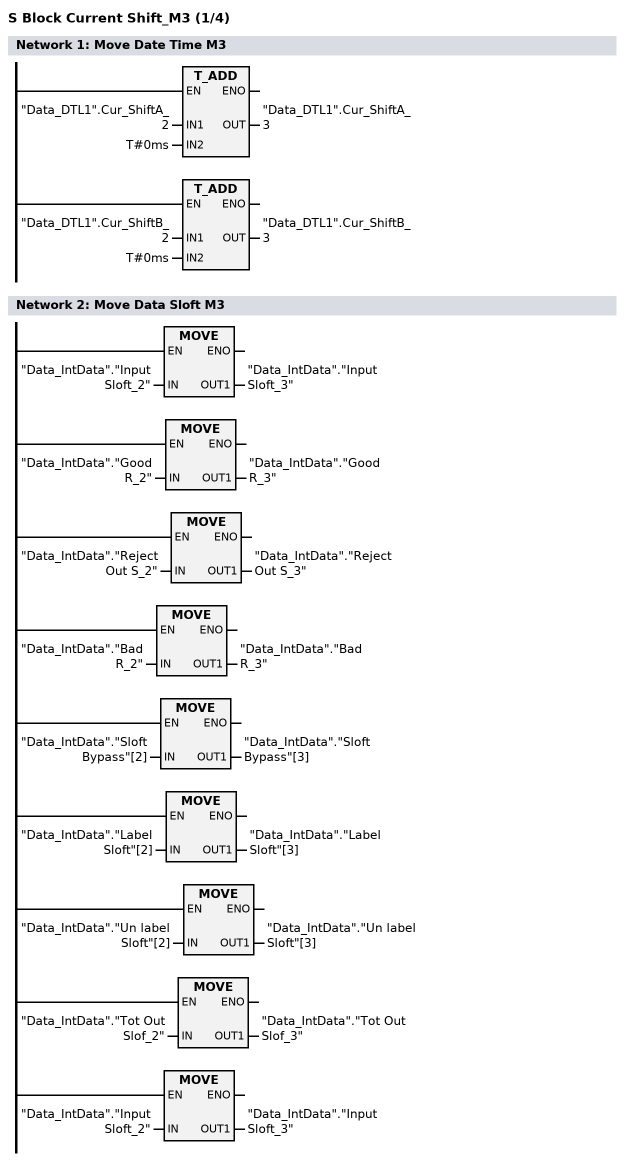
   "Data_DTL1".Cur_ShiftA_3 := T_ADD(IN1 := "Data_DTL1".Cur_ShiftA_2, IN2 := T#0ms);
   "Data_DTL1".Cur_ShiftB_3 := T_ADD(IN1 := "Data_DTL1".Cur_ShiftB_2, IN2 := T#0ms);
END_REGION

REGION Network 2: Move Data Sloft M3
   RUNG wire#powerrail
      { S7_GenerateENO := "TRUE" } Move(in := "Data_IntData"."Input Sloft_2", out1 => "Data_IntData"."Input Sloft_3")
   END_RUNG
   RUNG wire#powerrail
      { S7_GenerateENO := "TRUE" } Move(in := "Data_IntData"."Good R_2", out1 => "Data_IntData"."Good R_3")
   END_RUNG
   RUNG wire#powerrail
      { S7_GenerateENO := "TRUE" } Move(in := "Data_IntData"."Reject Out S_2", out1 => "Data_IntData"."Reject Out S_3")
   END_RUNG
   RUNG wire#powerrail
      { S7_GenerateENO := "TRUE" } Move(in := "Data_IntData"."Bad R_2", out1 => "Data_IntData"."Bad R_3")
   END_RUNG
   RUNG wire#powerrail
      { S7_GenerateENO := "TRUE" } Move(in := "Data_IntData"."Sloft Bypass"[2], out1 => "Data_IntData"."Sloft Bypass"[3])
   END_RUNG
   RUNG wire#powerrail
      { S7_GenerateENO := "TRUE" } Move(in := "Data_IntData"."Label Sloft"[2], out1 => "Data_IntData"."Label Sloft"[3])
   END_RUNG
   RUNG wire#powerrail
      { S7_GenerateENO := "TRUE" } Move(in := "Data_IntData"."Un label Sloft"[2], out1 => "Data_IntData"."Un label Sloft"[3])
   END_RUNG
   RUNG wire#powerrail
      { S7_GenerateENO := "TRUE" } Move(in := "Data_IntData"."Tot Out Slof_2", out1 => "Data_IntData"."Tot Out Slof_3")
   END_RUNG
   RUNG wire#powerrail
      { S7_GenerateENO := "TRUE" } Move(in := "Data_IntData"."Input Sloft_2", out1 => "Data_IntData"."Input Sloft_3")
   END_RUNG
   // the same network as SCL:
   "Data_IntData"."Input Sloft_3" := "Data_IntData"."Input Sloft_2";
   "Data_IntData"."Good R_3" := "Data_IntData"."Good R_2";
   "Data_IntData"."Reject Out S_3" := "Data_IntData"."Reject Out S_2";
   "Data_IntData"."Bad R_3" := "Data_IntData"."Bad R_2";
   "Data_IntData"."Sloft Bypass"[3] := "Data_IntData"."Sloft Bypass"[2];
   "Data_IntData"."Label Sloft"[3] := "Data_IntData"."Label Sloft"[2];
   "Data_IntData"."Un label Sloft"[3] := "Data_IntData"."Un label Sloft"[2];
   "Data_IntData"."Tot Out Slof_3" := "Data_IntData"."Tot Out Slof_2";
   "Data_IntData"."Input Sloft_3" := "Data_IntData"."Input Sloft_2";
END_REGION

REGION Network 3: Move Data Sloft Trigger & Aplicator M3
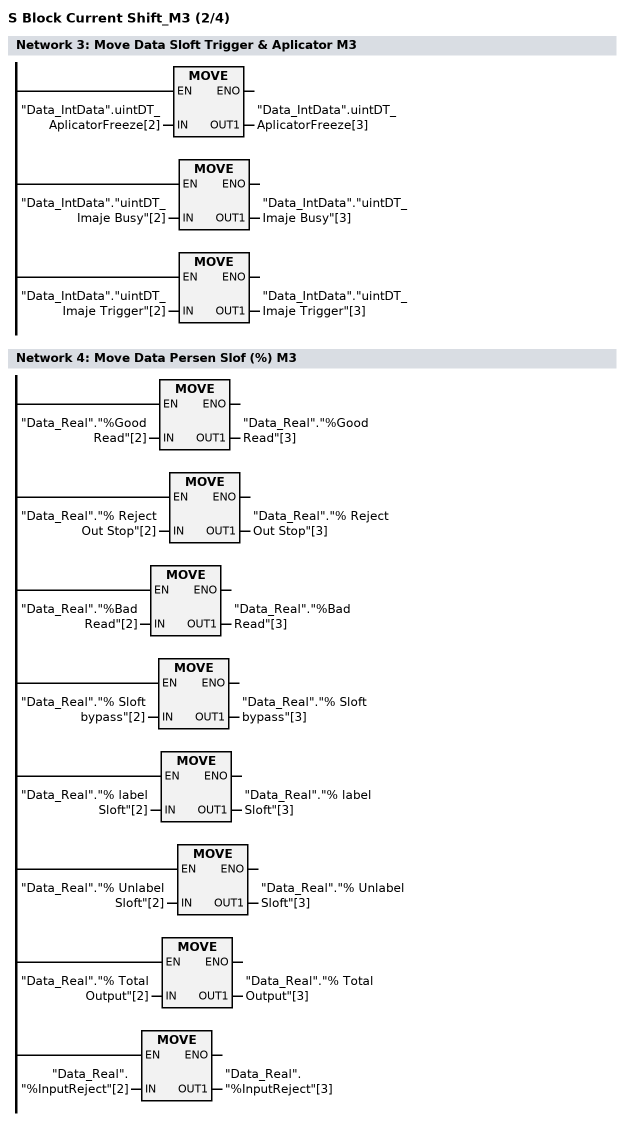
   RUNG wire#powerrail
      { S7_GenerateENO := "TRUE" } Move(in := "Data_IntData".uintDT_AplicatorFreeze[2], out1 => "Data_IntData".uintDT_AplicatorFreeze[3])
   END_RUNG
   RUNG wire#powerrail
      { S7_GenerateENO := "TRUE" } Move(in := "Data_IntData"."uintDT_Imaje Busy"[2], out1 => "Data_IntData"."uintDT_Imaje Busy"[3])
   END_RUNG
   RUNG wire#powerrail
      { S7_GenerateENO := "TRUE" } Move(in := "Data_IntData"."uintDT_Imaje Trigger"[2], out1 => "Data_IntData"."uintDT_Imaje Trigger"[3])
   END_RUNG
   // the same network as SCL:
   "Data_IntData".uintDT_AplicatorFreeze[3] := "Data_IntData".uintDT_AplicatorFreeze[2];
   "Data_IntData"."uintDT_Imaje Busy"[3] := "Data_IntData"."uintDT_Imaje Busy"[2];
   "Data_IntData"."uintDT_Imaje Trigger"[3] := "Data_IntData"."uintDT_Imaje Trigger"[2];
END_REGION

REGION Network 4: Move Data Persen Slof (%) M3
   RUNG wire#powerrail
      { S7_GenerateENO := "TRUE" } Move(in := "Data_Real"."%Good Read"[2], out1 => "Data_Real"."%Good Read"[3])
   END_RUNG
   RUNG wire#powerrail
      { S7_GenerateENO := "TRUE" } Move(in := "Data_Real"."% Reject Out Stop"[2], out1 => "Data_Real"."% Reject Out Stop"[3])
   END_RUNG
   RUNG wire#powerrail
      { S7_GenerateENO := "TRUE" } Move(in := "Data_Real"."%Bad Read"[2], out1 => "Data_Real"."%Bad Read"[3])
   END_RUNG
   RUNG wire#powerrail
      { S7_GenerateENO := "TRUE" } Move(in := "Data_Real"."% Sloft bypass"[2], out1 => "Data_Real"."% Sloft bypass"[3])
   END_RUNG
   RUNG wire#powerrail
      { S7_GenerateENO := "TRUE" } Move(in := "Data_Real"."% label Sloft"[2], out1 => "Data_Real"."% label Sloft"[3])
   END_RUNG
   RUNG wire#powerrail
      { S7_GenerateENO := "TRUE" } Move(in := "Data_Real"."% Unlabel Sloft"[2], out1 => "Data_Real"."% Unlabel Sloft"[3])
   END_RUNG
   RUNG wire#powerrail
      { S7_GenerateENO := "TRUE" } Move(in := "Data_Real"."% Total Output"[2], out1 => "Data_Real"."% Total Output"[3])
   END_RUNG
   RUNG wire#powerrail
      { S7_GenerateENO := "TRUE" } Move(in := "Data_Real"."%InputReject"[2], out1 => "Data_Real"."%InputReject"[3])
   END_RUNG
   // the same network as SCL:
   "Data_Real"."%Good Read"[3] := "Data_Real"."%Good Read"[2];
   "Data_Real"."% Reject Out Stop"[3] := "Data_Real"."% Reject Out Stop"[2];
   "Data_Real"."%Bad Read"[3] := "Data_Real"."%Bad Read"[2];
   "Data_Real"."% Sloft bypass"[3] := "Data_Real"."% Sloft bypass"[2];
   "Data_Real"."% label Sloft"[3] := "Data_Real"."% label Sloft"[2];
   "Data_Real"."% Unlabel Sloft"[3] := "Data_Real"."% Unlabel Sloft"[2];
   "Data_Real"."% Total Output"[3] := "Data_Real"."% Total Output"[2];
   "Data_Real"."%InputReject"[3] := "Data_Real"."%InputReject"[2];
END_REGION

REGION Network 5: Move Data Time Mesin M3
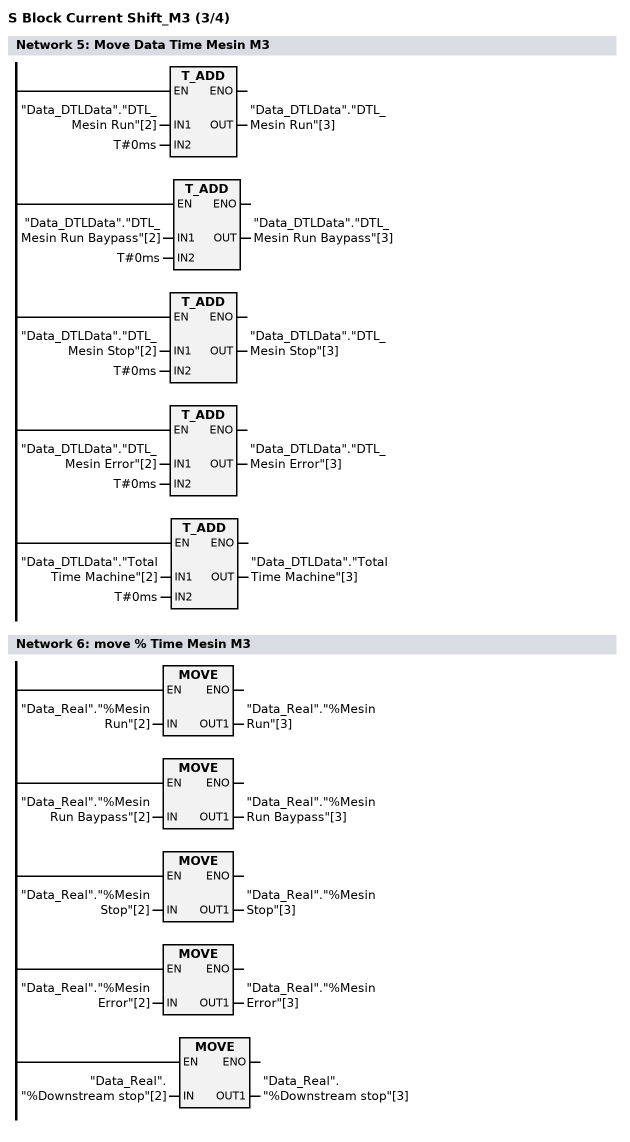
   "Data_DTLData"."DTL_Mesin Run"[3] := T_ADD(IN1 := "Data_DTLData"."DTL_Mesin Run"[2], IN2 := T#0ms);
   "Data_DTLData"."DTL_Mesin Run Baypass"[3] := T_ADD(IN1 := "Data_DTLData"."DTL_Mesin Run Baypass"[2],
                           IN2 := T#0ms);
   "Data_DTLData"."DTL_Mesin Stop"[3] := T_ADD(IN1 := "Data_DTLData"."DTL_Mesin Stop"[2], IN2 := T#0ms);
   "Data_DTLData"."DTL_Mesin Error"[3] := T_ADD(IN1 := "Data_DTLData"."DTL_Mesin Error"[2], IN2 := T#0ms);
   "Data_DTLData"."Total Time Machine"[3] := T_ADD(IN1 := "Data_DTLData"."Total Time Machine"[2], IN2 := T#0ms);
END_REGION

REGION Network 6: move % Time Mesin M3
   RUNG wire#powerrail
      { S7_GenerateENO := "TRUE" } Move(in := "Data_Real"."%Mesin Run"[2], out1 => "Data_Real"."%Mesin Run"[3])
   END_RUNG
   RUNG wire#powerrail
      { S7_GenerateENO := "TRUE" } Move(in := "Data_Real"."%Mesin Run Baypass"[2], out1 => "Data_Real"."%Mesin Run Baypass"[3])
   END_RUNG
   RUNG wire#powerrail
      { S7_GenerateENO := "TRUE" } Move(in := "Data_Real"."%Mesin Stop"[2], out1 => "Data_Real"."%Mesin Stop"[3])
   END_RUNG
   RUNG wire#powerrail
      { S7_GenerateENO := "TRUE" } Move(in := "Data_Real"."%Mesin Error"[2], out1 => "Data_Real"."%Mesin Error"[3])
   END_RUNG
   RUNG wire#powerrail
      { S7_GenerateENO := "TRUE" } Move(in := "Data_Real"."%Downstream stop"[2], out1 => "Data_Real"."%Downstream stop"[3])
   END_RUNG
   // the same network as SCL:
   "Data_Real"."%Mesin Run"[3] := "Data_Real"."%Mesin Run"[2];
   "Data_Real"."%Mesin Run Baypass"[3] := "Data_Real"."%Mesin Run Baypass"[2];
   "Data_Real"."%Mesin Stop"[3] := "Data_Real"."%Mesin Stop"[2];
   "Data_Real"."%Mesin Error"[3] := "Data_Real"."%Mesin Error"[2];
   "Data_Real"."%Downstream stop"[3] := "Data_Real"."%Downstream stop"[2];
END_REGION

REGION Network 7: Move Counter Error M3
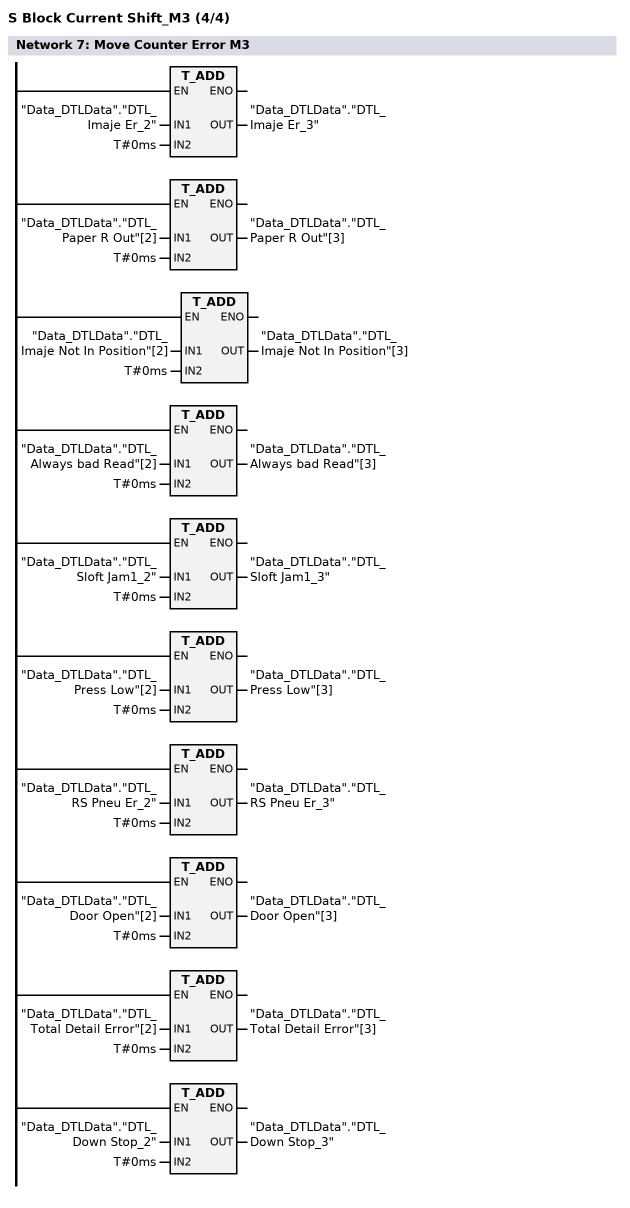
   "Data_DTLData"."DTL_Imaje Er_3" := T_ADD(IN1 := "Data_DTLData"."DTL_Imaje Er_2", IN2 := T#0ms);
   "Data_DTLData"."DTL_Paper R Out"[3] := T_ADD(IN1 := "Data_DTLData"."DTL_Paper R Out"[2], IN2 := T#0ms);
   "Data_DTLData"."DTL_Imaje Not In Position"[3] := T_ADD(IN1 := "Data_DTLData"."DTL_Imaje Not In Position"[2],
                           IN2 := T#0ms);
   "Data_DTLData"."DTL_Always bad Read"[3] := T_ADD(IN1 := "Data_DTLData"."DTL_Always bad Read"[2],
                           IN2 := T#0ms);
   "Data_DTLData"."DTL_Sloft Jam1_3" := T_ADD(IN1 := "Data_DTLData"."DTL_Sloft Jam1_2", IN2 := T#0ms);
   "Data_DTLData"."DTL_Press Low"[3] := T_ADD(IN1 := "Data_DTLData"."DTL_Press Low"[2], IN2 := T#0ms);
   "Data_DTLData"."DTL_RS Pneu Er_3" := T_ADD(IN1 := "Data_DTLData"."DTL_RS Pneu Er_2", IN2 := T#0ms);
   "Data_DTLData"."DTL_Door Open"[3] := T_ADD(IN1 := "Data_DTLData"."DTL_Door Open"[2], IN2 := T#0ms);
   "Data_DTLData"."DTL_Total Detail Error"[3] := T_ADD(IN1 := "Data_DTLData"."DTL_Total Detail Error"[2],
                           IN2 := T#0ms);
   "Data_DTLData"."DTL_Down Stop_3" := T_ADD(IN1 := "Data_DTLData"."DTL_Down Stop_2", IN2 := T#0ms);
END_REGION
END_FUNCTION_BLOCK

FUNCTION_BLOCK "S Block Current Shift_M4"   // FB13, LAD
{ S7_Optimized_Access := 'TRUE' }
VERSION : 0.1
BEGIN

REGION Network 1: Move Date Time M4
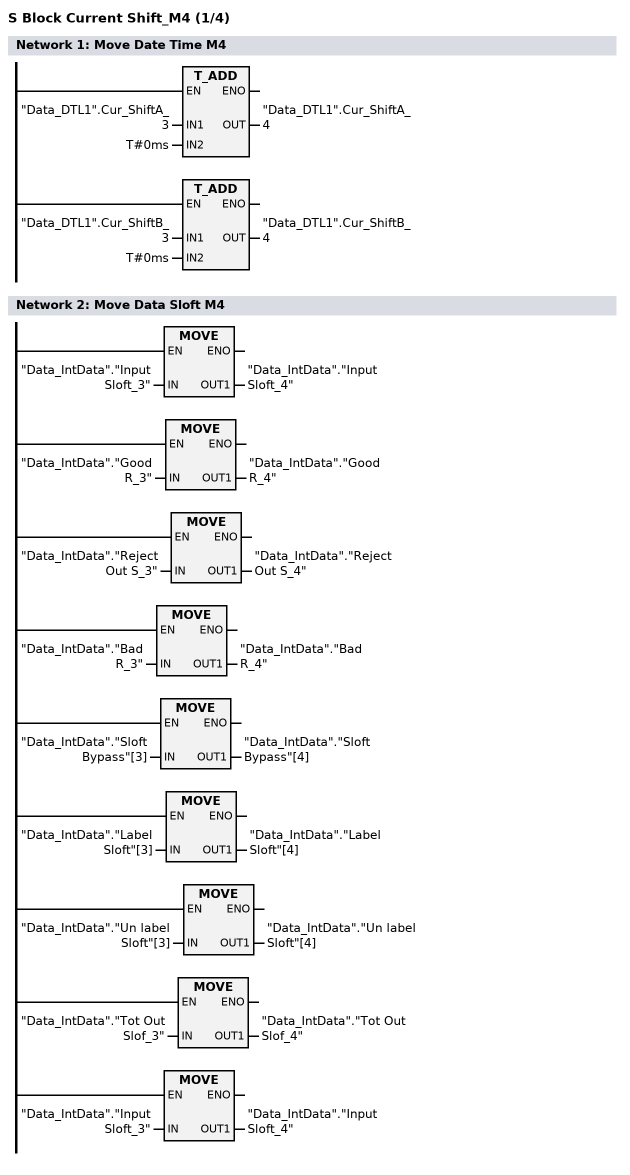
   "Data_DTL1".Cur_ShiftA_4 := T_ADD(IN1 := "Data_DTL1".Cur_ShiftA_3, IN2 := T#0ms);
   "Data_DTL1".Cur_ShiftB_4 := T_ADD(IN1 := "Data_DTL1".Cur_ShiftB_3, IN2 := T#0ms);
END_REGION

REGION Network 2: Move Data Sloft M4
   RUNG wire#powerrail
      { S7_GenerateENO := "TRUE" } Move(in := "Data_IntData"."Input Sloft_3", out1 => "Data_IntData"."Input Sloft_4")
   END_RUNG
   RUNG wire#powerrail
      { S7_GenerateENO := "TRUE" } Move(in := "Data_IntData"."Good R_3", out1 => "Data_IntData"."Good R_4")
   END_RUNG
   RUNG wire#powerrail
      { S7_GenerateENO := "TRUE" } Move(in := "Data_IntData"."Reject Out S_3", out1 => "Data_IntData"."Reject Out S_4")
   END_RUNG
   RUNG wire#powerrail
      { S7_GenerateENO := "TRUE" } Move(in := "Data_IntData"."Bad R_3", out1 => "Data_IntData"."Bad R_4")
   END_RUNG
   RUNG wire#powerrail
      { S7_GenerateENO := "TRUE" } Move(in := "Data_IntData"."Sloft Bypass"[3], out1 => "Data_IntData"."Sloft Bypass"[4])
   END_RUNG
   RUNG wire#powerrail
      { S7_GenerateENO := "TRUE" } Move(in := "Data_IntData"."Label Sloft"[3], out1 => "Data_IntData"."Label Sloft"[4])
   END_RUNG
   RUNG wire#powerrail
      { S7_GenerateENO := "TRUE" } Move(in := "Data_IntData"."Un label Sloft"[3], out1 => "Data_IntData"."Un label Sloft"[4])
   END_RUNG
   RUNG wire#powerrail
      { S7_GenerateENO := "TRUE" } Move(in := "Data_IntData"."Tot Out Slof_3", out1 => "Data_IntData"."Tot Out Slof_4")
   END_RUNG
   RUNG wire#powerrail
      { S7_GenerateENO := "TRUE" } Move(in := "Data_IntData"."Input Sloft_3", out1 => "Data_IntData"."Input Sloft_4")
   END_RUNG
   // the same network as SCL:
   "Data_IntData"."Input Sloft_4" := "Data_IntData"."Input Sloft_3";
   "Data_IntData"."Good R_4" := "Data_IntData"."Good R_3";
   "Data_IntData"."Reject Out S_4" := "Data_IntData"."Reject Out S_3";
   "Data_IntData"."Bad R_4" := "Data_IntData"."Bad R_3";
   "Data_IntData"."Sloft Bypass"[4] := "Data_IntData"."Sloft Bypass"[3];
   "Data_IntData"."Label Sloft"[4] := "Data_IntData"."Label Sloft"[3];
   "Data_IntData"."Un label Sloft"[4] := "Data_IntData"."Un label Sloft"[3];
   "Data_IntData"."Tot Out Slof_4" := "Data_IntData"."Tot Out Slof_3";
   "Data_IntData"."Input Sloft_4" := "Data_IntData"."Input Sloft_3";
END_REGION

REGION Network 3: Move Data Sloft Trigger & Aplicator M4
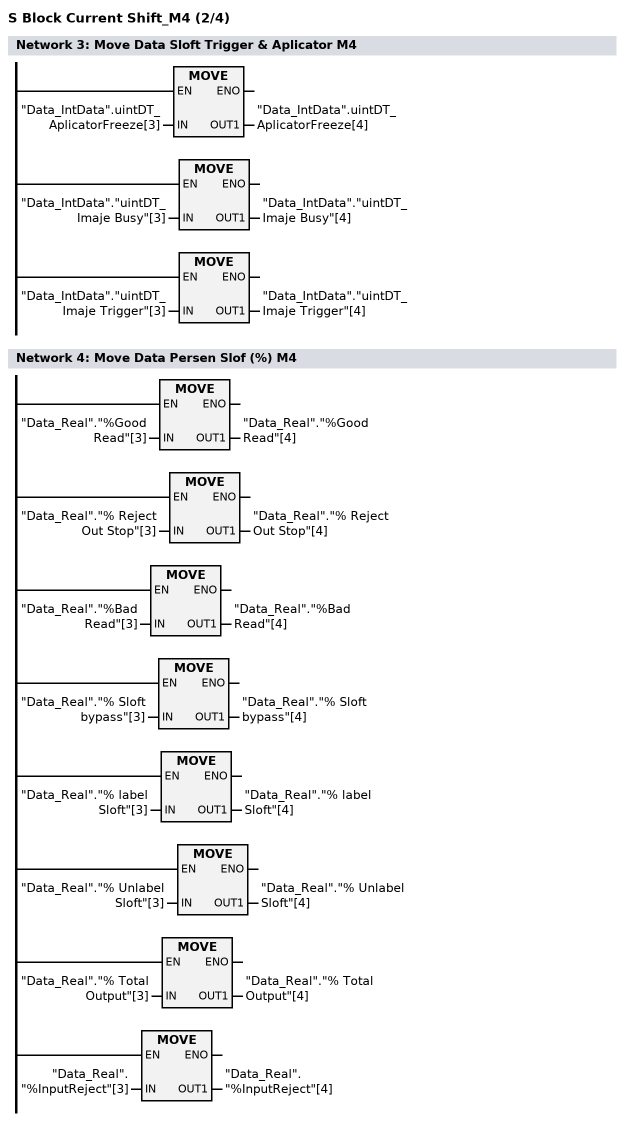
   RUNG wire#powerrail
      { S7_GenerateENO := "TRUE" } Move(in := "Data_IntData".uintDT_AplicatorFreeze[3], out1 => "Data_IntData".uintDT_AplicatorFreeze[4])
   END_RUNG
   RUNG wire#powerrail
      { S7_GenerateENO := "TRUE" } Move(in := "Data_IntData"."uintDT_Imaje Busy"[3], out1 => "Data_IntData"."uintDT_Imaje Busy"[4])
   END_RUNG
   RUNG wire#powerrail
      { S7_GenerateENO := "TRUE" } Move(in := "Data_IntData"."uintDT_Imaje Trigger"[3], out1 => "Data_IntData"."uintDT_Imaje Trigger"[4])
   END_RUNG
   // the same network as SCL:
   "Data_IntData".uintDT_AplicatorFreeze[4] := "Data_IntData".uintDT_AplicatorFreeze[3];
   "Data_IntData"."uintDT_Imaje Busy"[4] := "Data_IntData"."uintDT_Imaje Busy"[3];
   "Data_IntData"."uintDT_Imaje Trigger"[4] := "Data_IntData"."uintDT_Imaje Trigger"[3];
END_REGION

REGION Network 4: Move Data Persen Slof (%) M4
   RUNG wire#powerrail
      { S7_GenerateENO := "TRUE" } Move(in := "Data_Real"."%Good Read"[3], out1 => "Data_Real"."%Good Read"[4])
   END_RUNG
   RUNG wire#powerrail
      { S7_GenerateENO := "TRUE" } Move(in := "Data_Real"."% Reject Out Stop"[3], out1 => "Data_Real"."% Reject Out Stop"[4])
   END_RUNG
   RUNG wire#powerrail
      { S7_GenerateENO := "TRUE" } Move(in := "Data_Real"."%Bad Read"[3], out1 => "Data_Real"."%Bad Read"[4])
   END_RUNG
   RUNG wire#powerrail
      { S7_GenerateENO := "TRUE" } Move(in := "Data_Real"."% Sloft bypass"[3], out1 => "Data_Real"."% Sloft bypass"[4])
   END_RUNG
   RUNG wire#powerrail
      { S7_GenerateENO := "TRUE" } Move(in := "Data_Real"."% label Sloft"[3], out1 => "Data_Real"."% label Sloft"[4])
   END_RUNG
   RUNG wire#powerrail
      { S7_GenerateENO := "TRUE" } Move(in := "Data_Real"."% Unlabel Sloft"[3], out1 => "Data_Real"."% Unlabel Sloft"[4])
   END_RUNG
   RUNG wire#powerrail
      { S7_GenerateENO := "TRUE" } Move(in := "Data_Real"."% Total Output"[3], out1 => "Data_Real"."% Total Output"[4])
   END_RUNG
   RUNG wire#powerrail
      { S7_GenerateENO := "TRUE" } Move(in := "Data_Real"."%InputReject"[3], out1 => "Data_Real"."%InputReject"[4])
   END_RUNG
   // the same network as SCL:
   "Data_Real"."%Good Read"[4] := "Data_Real"."%Good Read"[3];
   "Data_Real"."% Reject Out Stop"[4] := "Data_Real"."% Reject Out Stop"[3];
   "Data_Real"."%Bad Read"[4] := "Data_Real"."%Bad Read"[3];
   "Data_Real"."% Sloft bypass"[4] := "Data_Real"."% Sloft bypass"[3];
   "Data_Real"."% label Sloft"[4] := "Data_Real"."% label Sloft"[3];
   "Data_Real"."% Unlabel Sloft"[4] := "Data_Real"."% Unlabel Sloft"[3];
   "Data_Real"."% Total Output"[4] := "Data_Real"."% Total Output"[3];
   "Data_Real"."%InputReject"[4] := "Data_Real"."%InputReject"[3];
END_REGION

REGION Network 5: Move Data Time Mesin M4
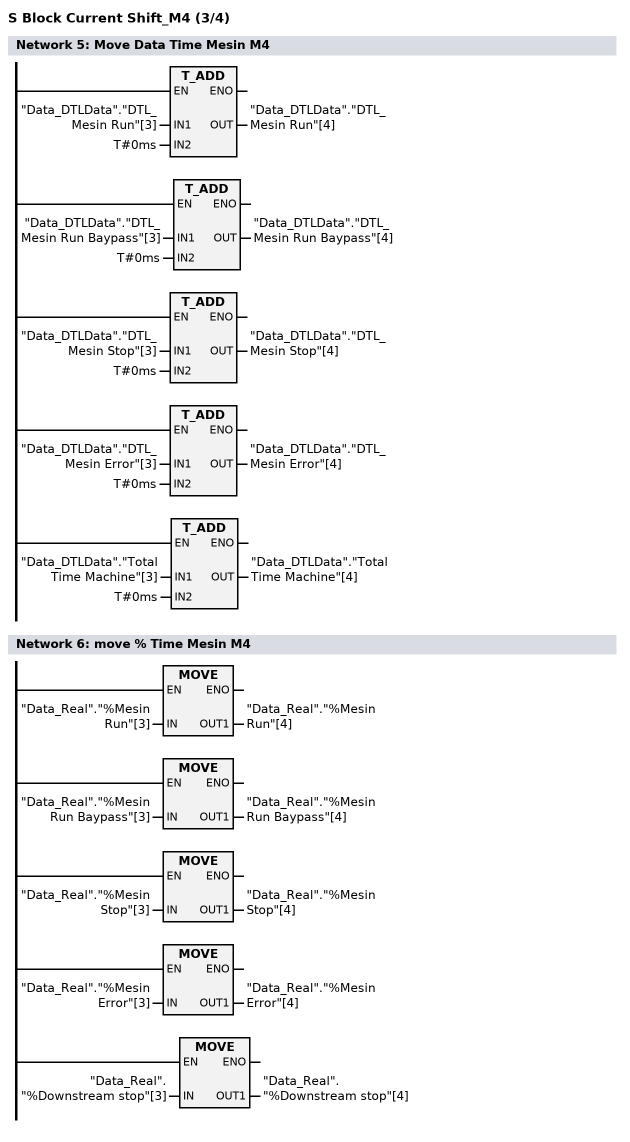
   "Data_DTLData"."DTL_Mesin Run"[4] := T_ADD(IN1 := "Data_DTLData"."DTL_Mesin Run"[3], IN2 := T#0ms);
   "Data_DTLData"."DTL_Mesin Run Baypass"[4] := T_ADD(IN1 := "Data_DTLData"."DTL_Mesin Run Baypass"[3],
                           IN2 := T#0ms);
   "Data_DTLData"."DTL_Mesin Stop"[4] := T_ADD(IN1 := "Data_DTLData"."DTL_Mesin Stop"[3], IN2 := T#0ms);
   "Data_DTLData"."DTL_Mesin Error"[4] := T_ADD(IN1 := "Data_DTLData"."DTL_Mesin Error"[3], IN2 := T#0ms);
   "Data_DTLData"."Total Time Machine"[4] := T_ADD(IN1 := "Data_DTLData"."Total Time Machine"[3], IN2 := T#0ms);
END_REGION

REGION Network 6: move % Time Mesin M4
   RUNG wire#powerrail
      { S7_GenerateENO := "TRUE" } Move(in := "Data_Real"."%Mesin Run"[3], out1 => "Data_Real"."%Mesin Run"[4])
   END_RUNG
   RUNG wire#powerrail
      { S7_GenerateENO := "TRUE" } Move(in := "Data_Real"."%Mesin Run Baypass"[3], out1 => "Data_Real"."%Mesin Run Baypass"[4])
   END_RUNG
   RUNG wire#powerrail
      { S7_GenerateENO := "TRUE" } Move(in := "Data_Real"."%Mesin Stop"[3], out1 => "Data_Real"."%Mesin Stop"[4])
   END_RUNG
   RUNG wire#powerrail
      { S7_GenerateENO := "TRUE" } Move(in := "Data_Real"."%Mesin Error"[3], out1 => "Data_Real"."%Mesin Error"[4])
   END_RUNG
   RUNG wire#powerrail
      { S7_GenerateENO := "TRUE" } Move(in := "Data_Real"."%Downstream stop"[3], out1 => "Data_Real"."%Downstream stop"[4])
   END_RUNG
   // the same network as SCL:
   "Data_Real"."%Mesin Run"[4] := "Data_Real"."%Mesin Run"[3];
   "Data_Real"."%Mesin Run Baypass"[4] := "Data_Real"."%Mesin Run Baypass"[3];
   "Data_Real"."%Mesin Stop"[4] := "Data_Real"."%Mesin Stop"[3];
   "Data_Real"."%Mesin Error"[4] := "Data_Real"."%Mesin Error"[3];
   "Data_Real"."%Downstream stop"[4] := "Data_Real"."%Downstream stop"[3];
END_REGION

REGION Network 7: Move Counter Error M4
